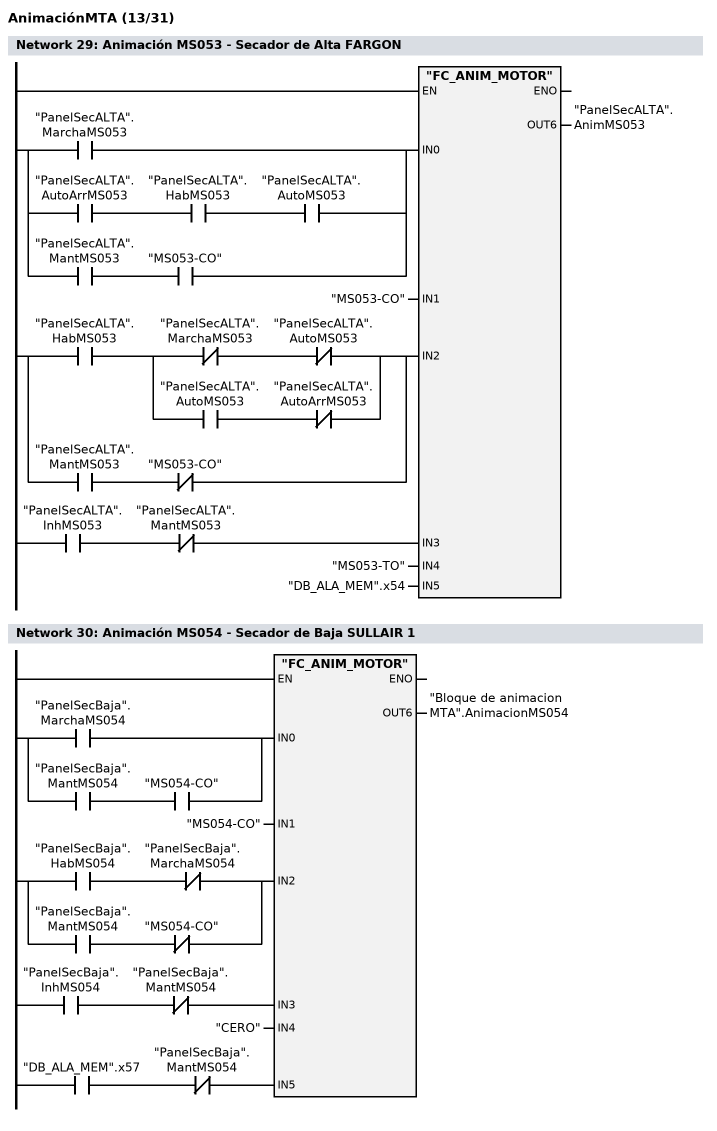
   RUNG wire#powerrail
      "FC_ANIM_MOTOR"(IN0 := wire#w1, IN2 := wire#w3, IN3 := wire#w4, IN1 := "MS053-CO", IN4 := "MS053-TO", IN5 := "DB_ALA_MEM".x54, OUT6 => "PanelSecALTA".AnimMS053)
   END_RUNG
   RUNG wire#powerrail
      Contact( "PanelSecALTA".MarchaMS053 )
   END_RUNG wire#w1
   RUNG wire#powerrail
      Contact( "PanelSecALTA".AutoArrMS053 )
      Contact( "PanelSecALTA".HabMS053 )
      Contact( "PanelSecALTA".AutoMS053 )
   END_RUNG wire#w1
   RUNG wire#powerrail
      Contact( "PanelSecALTA".MantMS053 )
      Contact( "MS053-CO" )
   END_RUNG wire#w1
   RUNG wire#powerrail
      Contact( "PanelSecALTA".HabMS053 )
      wire#w2
      I_Contact( "PanelSecALTA".MarchaMS053 )
      I_Contact( "PanelSecALTA".AutoMS053 )
   END_RUNG wire#w3
   RUNG wire#w2
      Contact( "PanelSecALTA".AutoMS053 )
      I_Contact( "PanelSecALTA".AutoArrMS053 )
   END_RUNG wire#w3
   RUNG wire#powerrail
      Contact( "PanelSecALTA".MantMS053 )
      I_Contact( "MS053-CO" )
   END_RUNG wire#w3
   RUNG wire#powerrail
      Contact( "PanelSecALTA".InhMS053 )
      I_Contact( "PanelSecALTA".MantMS053 )
   END_RUNG wire#w4
   // the same network as SCL:
   "FC_ANIM_MOTOR"(IN0 := "PanelSecALTA".MarchaMS053 OR ("PanelSecALTA".AutoArrMS053 AND "PanelSecALTA".HabMS053 AND "PanelSecALTA".AutoMS053) OR ("PanelSecALTA".MantMS053 AND "MS053-CO"),
                   IN1 := "MS053-CO",
                   IN2 := ("PanelSecALTA".HabMS053 AND ((NOT "PanelSecALTA".MarchaMS053 AND NOT "PanelSecALTA".AutoMS053) OR ("PanelSecALTA".AutoMS053 AND NOT "PanelSecALTA".AutoArrMS053))) OR ("PanelSecALTA".MantMS053 AND NOT "MS053-CO"),
                   IN3 := "PanelSecALTA".InhMS053 AND NOT "PanelSecALTA".MantMS053,
                   IN4 := "MS053-TO",
                   IN5 := "DB_ALA_MEM".x54,
                   OUT6 => "PanelSecALTA".AnimMS053);
END_REGION

REGION Network 30: Animación MS054 - Secador de Baja SULLAIR 1
   RUNG wire#powerrail
      "FC_ANIM_MOTOR"(IN0 := wire#w1, IN2 := wire#w2, IN3 := wire#w3, IN5 := wire#w4, IN1 := "MS054-CO", IN4 := "CERO", OUT6 => "Bloque de animacion MTA".AnimacionMS054)
   END_RUNG
   RUNG wire#powerrail
      Contact( "PanelSecBaja".MarchaMS054 )
   END_RUNG wire#w1
   RUNG wire#powerrail
      Contact( "PanelSecBaja".MantMS054 )
      Contact( "MS054-CO" )
   END_RUNG wire#w1
   RUNG wire#powerrail
      Contact( "PanelSecBaja".HabMS054 )
      I_Contact( "PanelSecBaja".MarchaMS054 )
   END_RUNG wire#w2
   RUNG wire#powerrail
      Contact( "PanelSecBaja".MantMS054 )
      I_Contact( "MS054-CO" )
   END_RUNG wire#w2
   RUNG wire#powerrail
      Contact( "PanelSecBaja".InhMS054 )
      I_Contact( "PanelSecBaja".MantMS054 )
   END_RUNG wire#w3
   RUNG wire#powerrail
      Contact( "DB_ALA_MEM".x57 )
      I_Contact( "PanelSecBaja".MantMS054 )
   END_RUNG wire#w4
   // the same network as SCL:
   "FC_ANIM_MOTOR"(IN0 := "PanelSecBaja".MarchaMS054 OR ("PanelSecBaja".MantMS054 AND "MS054-CO"),
                   IN1 := "MS054-CO",
                   IN2 := ("PanelSecBaja".HabMS054 AND NOT "PanelSecBaja".MarchaMS054) OR ("PanelSecBaja".MantMS054 AND NOT "MS054-CO"),
                   IN3 := "PanelSecBaja".InhMS054 AND NOT "PanelSecBaja".MantMS054,
                   IN4 := "CERO",
                   IN5 := "DB_ALA_MEM".x57 AND NOT "PanelSecBaja".MantMS054,
                   OUT6 => "Bloque de animacion MTA".AnimacionMS054);
END_REGION

REGION Network 31: Animación MS055 - Secador de Baja SULLAIR 2
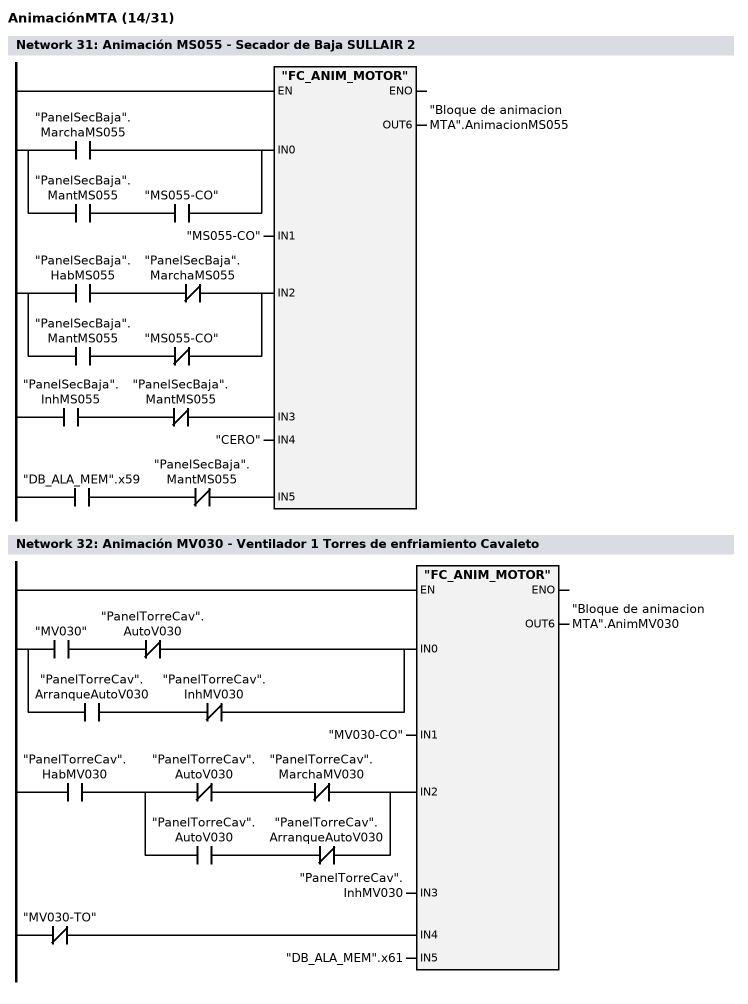
   RUNG wire#powerrail
      "FC_ANIM_MOTOR"(IN0 := wire#w1, IN2 := wire#w2, IN3 := wire#w3, IN5 := wire#w4, IN1 := "MS055-CO", IN4 := "CERO", OUT6 => "Bloque de animacion MTA".AnimacionMS055)
   END_RUNG
   RUNG wire#powerrail
      Contact( "PanelSecBaja".MarchaMS055 )
   END_RUNG wire#w1
   RUNG wire#powerrail
      Contact( "PanelSecBaja".MantMS055 )
      Contact( "MS055-CO" )
   END_RUNG wire#w1
   RUNG wire#powerrail
      Contact( "PanelSecBaja".HabMS055 )
      I_Contact( "PanelSecBaja".MarchaMS055 )
   END_RUNG wire#w2
   RUNG wire#powerrail
      Contact( "PanelSecBaja".MantMS055 )
      I_Contact( "MS055-CO" )
   END_RUNG wire#w2
   RUNG wire#powerrail
      Contact( "PanelSecBaja".InhMS055 )
      I_Contact( "PanelSecBaja".MantMS055 )
   END_RUNG wire#w3
   RUNG wire#powerrail
      Contact( "DB_ALA_MEM".x59 )
      I_Contact( "PanelSecBaja".MantMS055 )
   END_RUNG wire#w4
   // the same network as SCL:
   "FC_ANIM_MOTOR"(IN0 := "PanelSecBaja".MarchaMS055 OR ("PanelSecBaja".MantMS055 AND "MS055-CO"),
                   IN1 := "MS055-CO",
                   IN2 := ("PanelSecBaja".HabMS055 AND NOT "PanelSecBaja".MarchaMS055) OR ("PanelSecBaja".MantMS055 AND NOT "MS055-CO"),
                   IN3 := "PanelSecBaja".InhMS055 AND NOT "PanelSecBaja".MantMS055,
                   IN4 := "CERO",
                   IN5 := "DB_ALA_MEM".x59 AND NOT "PanelSecBaja".MantMS055,
                   OUT6 => "Bloque de animacion MTA".AnimacionMS055);
END_REGION

REGION Network 32: Animación MV030 - Ventilador 1 Torres de enfriamiento Cavaleto
   RUNG wire#powerrail
      "FC_ANIM_MOTOR"(IN0 := wire#w1, IN2 := wire#w3, IN4 := wire#w4, IN1 := "MV030-CO", IN3 := "PanelTorreCav".InhMV030, IN5 := "DB_ALA_MEM".x61, OUT6 => "Bloque de animacion MTA".AnimMV030)
   END_RUNG
   RUNG wire#powerrail
      Contact( "MV030" )
      I_Contact( "PanelTorreCav".AutoV030 )
   END_RUNG wire#w1
   RUNG wire#powerrail
      Contact( "PanelTorreCav".ArranqueAutoV030 )
      I_Contact( "PanelTorreCav".InhMV030 )
   END_RUNG wire#w1
   RUNG wire#powerrail
      Contact( "PanelTorreCav".HabMV030 )
      wire#w2
      I_Contact( "PanelTorreCav".AutoV030 )
      I_Contact( "PanelTorreCav".MarchaMV030 )
   END_RUNG wire#w3
   RUNG wire#w2
      Contact( "PanelTorreCav".AutoV030 )
      I_Contact( "PanelTorreCav".ArranqueAutoV030 )
   END_RUNG wire#w3
   RUNG wire#powerrail
      I_Contact( "MV030-TO" )
   END_RUNG wire#w4
   // the same network as SCL:
   "FC_ANIM_MOTOR"(IN0 := ("MV030" AND NOT "PanelTorreCav".AutoV030) OR ("PanelTorreCav".ArranqueAutoV030 AND NOT "PanelTorreCav".InhMV030),
                   IN1 := "MV030-CO",
                   IN2 := "PanelTorreCav".HabMV030 AND ((NOT "PanelTorreCav".AutoV030 AND NOT "PanelTorreCav".MarchaMV030) OR ("PanelTorreCav".AutoV030 AND NOT "PanelTorreCav".ArranqueAutoV030)),
                   IN3 := "PanelTorreCav".InhMV030,
                   IN4 := NOT "MV030-TO",
                   IN5 := "DB_ALA_MEM".x61,
                   OUT6 => "Bloque de animacion MTA".AnimMV030);
END_REGION

REGION Network 33: Animación MV031 - Ventilador 2 Torres de enfriamiento Cavaleto
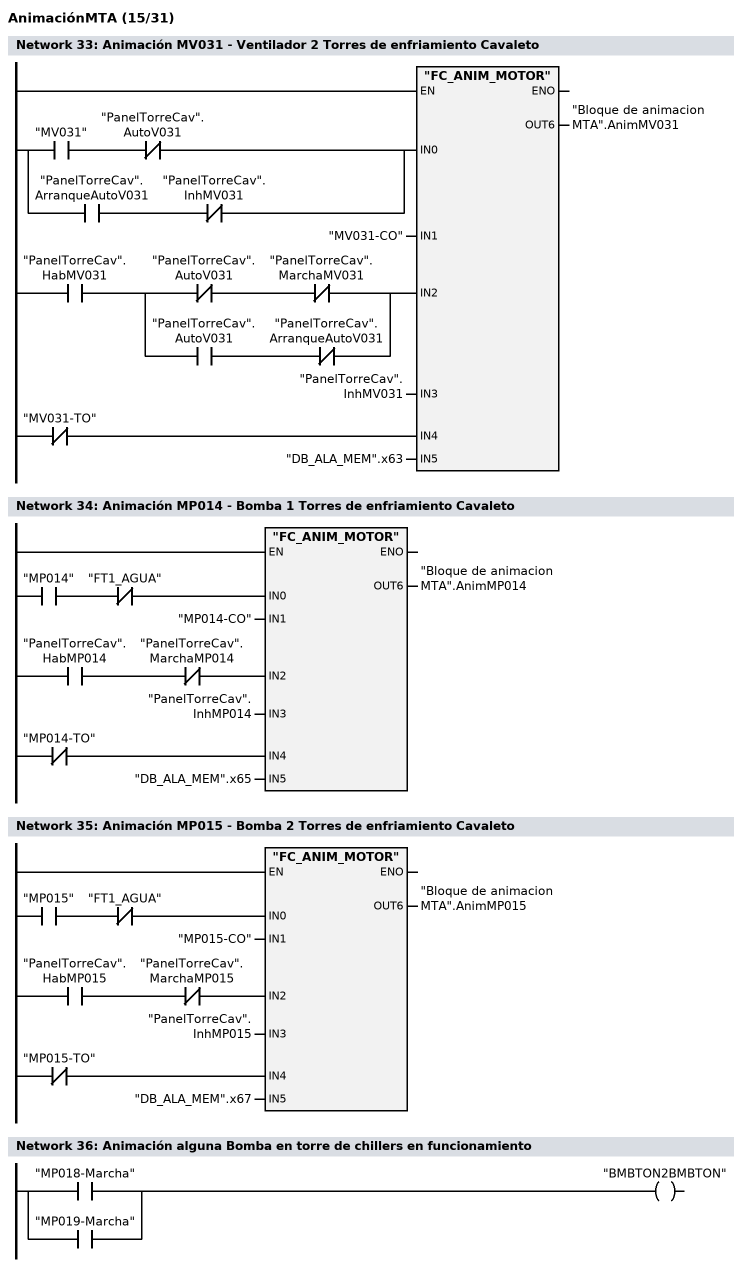
   RUNG wire#powerrail
      "FC_ANIM_MOTOR"(IN0 := wire#w1, IN2 := wire#w3, IN4 := wire#w4, IN1 := "MV031-CO", IN3 := "PanelTorreCav".InhMV031, IN5 := "DB_ALA_MEM".x63, OUT6 => "Bloque de animacion MTA".AnimMV031)
   END_RUNG
   RUNG wire#powerrail
      Contact( "MV031" )
      I_Contact( "PanelTorreCav".AutoV031 )
   END_RUNG wire#w1
   RUNG wire#powerrail
      Contact( "PanelTorreCav".ArranqueAutoV031 )
      I_Contact( "PanelTorreCav".InhMV031 )
   END_RUNG wire#w1
   RUNG wire#powerrail
      Contact( "PanelTorreCav".HabMV031 )
      wire#w2
      I_Contact( "PanelTorreCav".AutoV031 )
      I_Contact( "PanelTorreCav".MarchaMV031 )
   END_RUNG wire#w3
   RUNG wire#w2
      Contact( "PanelTorreCav".AutoV031 )
      I_Contact( "PanelTorreCav".ArranqueAutoV031 )
   END_RUNG wire#w3
   RUNG wire#powerrail
      I_Contact( "MV031-TO" )
   END_RUNG wire#w4
   // the same network as SCL:
   "FC_ANIM_MOTOR"(IN0 := ("MV031" AND NOT "PanelTorreCav".AutoV031) OR ("PanelTorreCav".ArranqueAutoV031 AND NOT "PanelTorreCav".InhMV031),
                   IN1 := "MV031-CO",
                   IN2 := "PanelTorreCav".HabMV031 AND ((NOT "PanelTorreCav".AutoV031 AND NOT "PanelTorreCav".MarchaMV031) OR ("PanelTorreCav".AutoV031 AND NOT "PanelTorreCav".ArranqueAutoV031)),
                   IN3 := "PanelTorreCav".InhMV031,
                   IN4 := NOT "MV031-TO",
                   IN5 := "DB_ALA_MEM".x63,
                   OUT6 => "Bloque de animacion MTA".AnimMV031);
END_REGION

REGION Network 34: Animación MP014 - Bomba 1 Torres de enfriamiento Cavaleto
   RUNG wire#powerrail
      "FC_ANIM_MOTOR"(IN0 := wire#w1, IN2 := wire#w2, IN4 := wire#w3, IN1 := "MP014-CO", IN3 := "PanelTorreCav".InhMP014, IN5 := "DB_ALA_MEM".x65, OUT6 => "Bloque de animacion MTA".AnimMP014)
   END_RUNG
   RUNG wire#powerrail
      Contact( "MP014" )
      I_Contact( "FT1_AGUA" )
   END_RUNG wire#w1
   RUNG wire#powerrail
      Contact( "PanelTorreCav".HabMP014 )
      I_Contact( "PanelTorreCav".MarchaMP014 )
   END_RUNG wire#w2
   RUNG wire#powerrail
      I_Contact( "MP014-TO" )
   END_RUNG wire#w3
   // the same network as SCL:
   "FC_ANIM_MOTOR"(IN0 := "MP014" AND NOT "FT1_AGUA",
                   IN1 := "MP014-CO",
                   IN2 := "PanelTorreCav".HabMP014 AND NOT "PanelTorreCav".MarchaMP014,
                   IN3 := "PanelTorreCav".InhMP014,
                   IN4 := NOT "MP014-TO",
                   IN5 := "DB_ALA_MEM".x65,
                   OUT6 => "Bloque de animacion MTA".AnimMP014);
END_REGION

REGION Network 35: Animación MP015 - Bomba 2 Torres de enfriamiento Cavaleto
   RUNG wire#powerrail
      "FC_ANIM_MOTOR"(IN0 := wire#w1, IN2 := wire#w2, IN4 := wire#w3, IN1 := "MP015-CO", IN3 := "PanelTorreCav".InhMP015, IN5 := "DB_ALA_MEM".x67, OUT6 => "Bloque de animacion MTA".AnimMP015)
   END_RUNG
   RUNG wire#powerrail
      Contact( "MP015" )
      I_Contact( "FT1_AGUA" )
   END_RUNG wire#w1
   RUNG wire#powerrail
      Contact( "PanelTorreCav".HabMP015 )
      I_Contact( "PanelTorreCav".MarchaMP015 )
   END_RUNG wire#w2
   RUNG wire#powerrail
      I_Contact( "MP015-TO" )
   END_RUNG wire#w3
   // the same network as SCL:
   "FC_ANIM_MOTOR"(IN0 := "MP015" AND NOT "FT1_AGUA",
                   IN1 := "MP015-CO",
                   IN2 := "PanelTorreCav".HabMP015 AND NOT "PanelTorreCav".MarchaMP015,
                   IN3 := "PanelTorreCav".InhMP015,
                   IN4 := NOT "MP015-TO",
                   IN5 := "DB_ALA_MEM".x67,
                   OUT6 => "Bloque de animacion MTA".AnimMP015);
END_REGION

REGION Network 36: Animación alguna Bomba en torre de chillers en funcionamiento
   RUNG wire#powerrail
      Contact( "MP018-Marcha" )
      wire#w1
      Coil( "BMBTON2BMBTON" )
   END_RUNG
   RUNG wire#powerrail
      Contact( "MP019-Marcha" )
   END_RUNG wire#w1
   // the same network as SCL:
   "BMBTON2BMBTON" := "MP018-Marcha" OR "MP019-Marcha";
END_REGION

REGION Network 37: Animación alguna Bomba en torre de cavaleto en funcionamiento
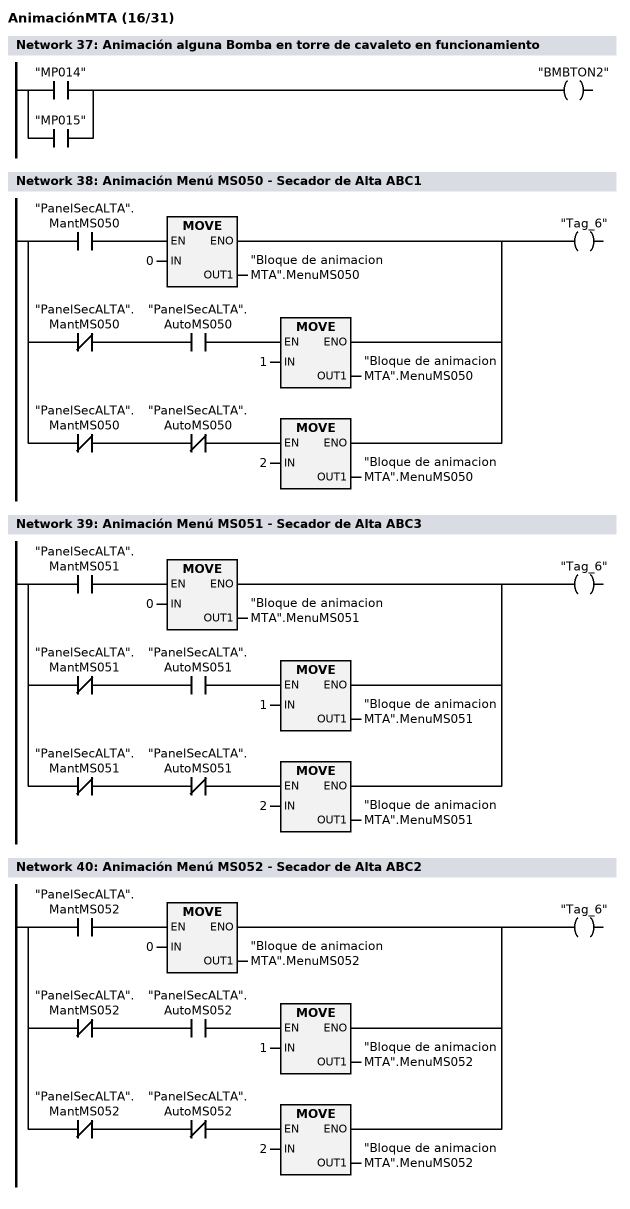
   RUNG wire#powerrail
      Contact( "MP014" )
      wire#w1
      Coil( "BMBTON2" )
   END_RUNG
   RUNG wire#powerrail
      Contact( "MP015" )
   END_RUNG wire#w1
   // the same network as SCL:
   "BMBTON2" := "MP014" OR "MP015";
END_REGION

REGION Network 38: Animación Menú MS050 - Secador de Alta ABC1
   RUNG wire#powerrail
      Contact( "PanelSecALTA".MantMS050 )
      { S7_GenerateENO := "TRUE" } Move(in := 0, out1 => "Bloque de animacion MTA".MenuMS050)
      wire#w1
      Coil( "Tag_6" )
   END_RUNG
   RUNG wire#powerrail
      I_Contact( "PanelSecALTA".MantMS050 )
      Contact( "PanelSecALTA".AutoMS050 )
      { S7_GenerateENO := "TRUE" } Move(in := 1, out1 => "Bloque de animacion MTA".MenuMS050)
   END_RUNG wire#w1
   RUNG wire#powerrail
      I_Contact( "PanelSecALTA".MantMS050 )
      I_Contact( "PanelSecALTA".AutoMS050 )
      { S7_GenerateENO := "TRUE" } Move(in := 2, out1 => "Bloque de animacion MTA".MenuMS050)
   END_RUNG wire#w1
   // the same network as SCL:
   // ENO of a box is taken as its EN; it also drops when the box reports an error
   IF "PanelSecALTA".MantMS050 THEN "Bloque de animacion MTA".MenuMS050 := 0; END_IF;
   #_w1 := NOT "PanelSecALTA".MantMS050 AND "PanelSecALTA".AutoMS050;
   IF #_w1 THEN "Bloque de animacion MTA".MenuMS050 := 1; END_IF;
   #_w2 := NOT "PanelSecALTA".MantMS050 AND NOT "PanelSecALTA".AutoMS050;
   IF #_w2 THEN "Bloque de animacion MTA".MenuMS050 := 2; END_IF;
   "Tag_6" := "PanelSecALTA".MantMS050 OR #_w1 OR #_w2;
END_REGION

REGION Network 39: Animación Menú MS051 - Secador de Alta ABC3
   RUNG wire#powerrail
      Contact( "PanelSecALTA".MantMS051 )
      { S7_GenerateENO := "TRUE" } Move(in := 0, out1 => "Bloque de animacion MTA".MenuMS051)
      wire#w1
      Coil( "Tag_6" )
   END_RUNG
   RUNG wire#powerrail
      I_Contact( "PanelSecALTA".MantMS051 )
      Contact( "PanelSecALTA".AutoMS051 )
      { S7_GenerateENO := "TRUE" } Move(in := 1, out1 => "Bloque de animacion MTA".MenuMS051)
   END_RUNG wire#w1
   RUNG wire#powerrail
      I_Contact( "PanelSecALTA".MantMS051 )
      I_Contact( "PanelSecALTA".AutoMS051 )
      { S7_GenerateENO := "TRUE" } Move(in := 2, out1 => "Bloque de animacion MTA".MenuMS051)
   END_RUNG wire#w1
   // the same network as SCL:
   // ENO of a box is taken as its EN; it also drops when the box reports an error
   IF "PanelSecALTA".MantMS051 THEN "Bloque de animacion MTA".MenuMS051 := 0; END_IF;
   #_w1 := NOT "PanelSecALTA".MantMS051 AND "PanelSecALTA".AutoMS051;
   IF #_w1 THEN "Bloque de animacion MTA".MenuMS051 := 1; END_IF;
   #_w2 := NOT "PanelSecALTA".MantMS051 AND NOT "PanelSecALTA".AutoMS051;
   IF #_w2 THEN "Bloque de animacion MTA".MenuMS051 := 2; END_IF;
   "Tag_6" := "PanelSecALTA".MantMS051 OR #_w1 OR #_w2;
END_REGION

REGION Network 40: Animación Menú MS052 - Secador de Alta ABC2
   RUNG wire#powerrail
      Contact( "PanelSecALTA".MantMS052 )
      { S7_GenerateENO := "TRUE" } Move(in := 0, out1 => "Bloque de animacion MTA".MenuMS052)
      wire#w1
      Coil( "Tag_6" )
   END_RUNG
   RUNG wire#powerrail
      I_Contact( "PanelSecALTA".MantMS052 )
      Contact( "PanelSecALTA".AutoMS052 )
      { S7_GenerateENO := "TRUE" } Move(in := 1, out1 => "Bloque de animacion MTA".MenuMS052)
   END_RUNG wire#w1
   RUNG wire#powerrail
      I_Contact( "PanelSecALTA".MantMS052 )
      I_Contact( "PanelSecALTA".AutoMS052 )
      { S7_GenerateENO := "TRUE" } Move(in := 2, out1 => "Bloque de animacion MTA".MenuMS052)
   END_RUNG wire#w1
   // the same network as SCL:
   // ENO of a box is taken as its EN; it also drops when the box reports an error
   IF "PanelSecALTA".MantMS052 THEN "Bloque de animacion MTA".MenuMS052 := 0; END_IF;
   #_w1 := NOT "PanelSecALTA".MantMS052 AND "PanelSecALTA".AutoMS052;
   IF #_w1 THEN "Bloque de animacion MTA".MenuMS052 := 1; END_IF;
   #_w2 := NOT "PanelSecALTA".MantMS052 AND NOT "PanelSecALTA".AutoMS052;
   IF #_w2 THEN "Bloque de animacion MTA".MenuMS052 := 2; END_IF;
   "Tag_6" := "PanelSecALTA".MantMS052 OR #_w1 OR #_w2;
END_REGION

REGION Network 41: Animación Menú MS053 - Secador de Alta FARGON
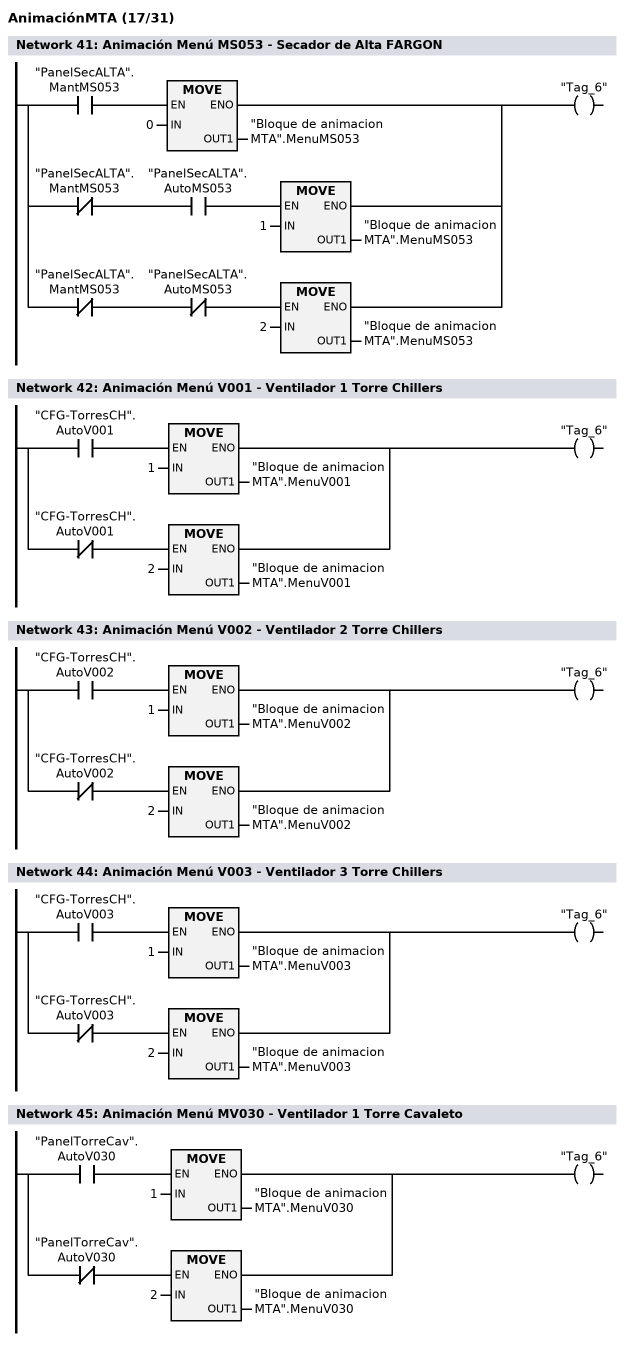
   RUNG wire#powerrail
      Contact( "PanelSecALTA".MantMS053 )
      { S7_GenerateENO := "TRUE" } Move(in := 0, out1 => "Bloque de animacion MTA".MenuMS053)
      wire#w1
      Coil( "Tag_6" )
   END_RUNG
   RUNG wire#powerrail
      I_Contact( "PanelSecALTA".MantMS053 )
      Contact( "PanelSecALTA".AutoMS053 )
      { S7_GenerateENO := "TRUE" } Move(in := 1, out1 => "Bloque de animacion MTA".MenuMS053)
   END_RUNG wire#w1
   RUNG wire#powerrail
      I_Contact( "PanelSecALTA".MantMS053 )
      I_Contact( "PanelSecALTA".AutoMS053 )
      { S7_GenerateENO := "TRUE" } Move(in := 2, out1 => "Bloque de animacion MTA".MenuMS053)
   END_RUNG wire#w1
   // the same network as SCL:
   // ENO of a box is taken as its EN; it also drops when the box reports an error
   IF "PanelSecALTA".MantMS053 THEN "Bloque de animacion MTA".MenuMS053 := 0; END_IF;
   #_w1 := NOT "PanelSecALTA".MantMS053 AND "PanelSecALTA".AutoMS053;
   IF #_w1 THEN "Bloque de animacion MTA".MenuMS053 := 1; END_IF;
   #_w2 := NOT "PanelSecALTA".MantMS053 AND NOT "PanelSecALTA".AutoMS053;
   IF #_w2 THEN "Bloque de animacion MTA".MenuMS053 := 2; END_IF;
   "Tag_6" := "PanelSecALTA".MantMS053 OR #_w1 OR #_w2;
END_REGION

REGION Network 42: Animación Menú V001 - Ventilador 1 Torre Chillers
   RUNG wire#powerrail
      Contact( "CFG-TorresCH".AutoV001 )
      { S7_GenerateENO := "TRUE" } Move(in := 1, out1 => "Bloque de animacion MTA".MenuV001)
      wire#w1
      Coil( "Tag_6" )
   END_RUNG
   RUNG wire#powerrail
      I_Contact( "CFG-TorresCH".AutoV001 )
      { S7_GenerateENO := "TRUE" } Move(in := 2, out1 => "Bloque de animacion MTA".MenuV001)
   END_RUNG wire#w1
   // the same network as SCL:
   // ENO of a box is taken as its EN; it also drops when the box reports an error
   IF "CFG-TorresCH".AutoV001 THEN "Bloque de animacion MTA".MenuV001 := 1; END_IF;
   #_w1 := NOT "CFG-TorresCH".AutoV001;
   IF #_w1 THEN "Bloque de animacion MTA".MenuV001 := 2; END_IF;
   "Tag_6" := "CFG-TorresCH".AutoV001 OR #_w1;
END_REGION

REGION Network 43: Animación Menú V002 - Ventilador 2 Torre Chillers
   RUNG wire#powerrail
      Contact( "CFG-TorresCH".AutoV002 )
      { S7_GenerateENO := "TRUE" } Move(in := 1, out1 => "Bloque de animacion MTA".MenuV002)
      wire#w1
      Coil( "Tag_6" )
   END_RUNG
   RUNG wire#powerrail
      I_Contact( "CFG-TorresCH".AutoV002 )
      { S7_GenerateENO := "TRUE" } Move(in := 2, out1 => "Bloque de animacion MTA".MenuV002)
   END_RUNG wire#w1
   // the same network as SCL:
   // ENO of a box is taken as its EN; it also drops when the box reports an error
   IF "CFG-TorresCH".AutoV002 THEN "Bloque de animacion MTA".MenuV002 := 1; END_IF;
   #_w1 := NOT "CFG-TorresCH".AutoV002;
   IF #_w1 THEN "Bloque de animacion MTA".MenuV002 := 2; END_IF;
   "Tag_6" := "CFG-TorresCH".AutoV002 OR #_w1;
END_REGION

REGION Network 44: Animación Menú V003 - Ventilador 3 Torre Chillers
   RUNG wire#powerrail
      Contact( "CFG-TorresCH".AutoV003 )
      { S7_GenerateENO := "TRUE" } Move(in := 1, out1 => "Bloque de animacion MTA".MenuV003)
      wire#w1
      Coil( "Tag_6" )
   END_RUNG
   RUNG wire#powerrail
      I_Contact( "CFG-TorresCH".AutoV003 )
      { S7_GenerateENO := "TRUE" } Move(in := 2, out1 => "Bloque de animacion MTA".MenuV003)
   END_RUNG wire#w1
   // the same network as SCL:
   // ENO of a box is taken as its EN; it also drops when the box reports an error
   IF "CFG-TorresCH".AutoV003 THEN "Bloque de animacion MTA".MenuV003 := 1; END_IF;
   #_w1 := NOT "CFG-TorresCH".AutoV003;
   IF #_w1 THEN "Bloque de animacion MTA".MenuV003 := 2; END_IF;
   "Tag_6" := "CFG-TorresCH".AutoV003 OR #_w1;
END_REGION

REGION Network 45: Animación Menú MV030 - Ventilador 1 Torre Cavaleto
   RUNG wire#powerrail
      Contact( "PanelTorreCav".AutoV030 )
      { S7_GenerateENO := "TRUE" } Move(in := 1, out1 => "Bloque de animacion MTA".MenuV030)
      wire#w1
      Coil( "Tag_6" )
   END_RUNG
   RUNG wire#powerrail
      I_Contact( "PanelTorreCav".AutoV030 )
      { S7_GenerateENO := "TRUE" } Move(in := 2, out1 => "Bloque de animacion MTA".MenuV030)
   END_RUNG wire#w1
   // the same network as SCL:
   // ENO of a box is taken as its EN; it also drops when the box reports an error
   IF "PanelTorreCav".AutoV030 THEN "Bloque de animacion MTA".MenuV030 := 1; END_IF;
   #_w1 := NOT "PanelTorreCav".AutoV030;
   IF #_w1 THEN "Bloque de animacion MTA".MenuV030 := 2; END_IF;
   "Tag_6" := "PanelTorreCav".AutoV030 OR #_w1;
END_REGION

REGION Network 46: Animación Menú MV031 - Ventilador 2 Torre Cavaleto
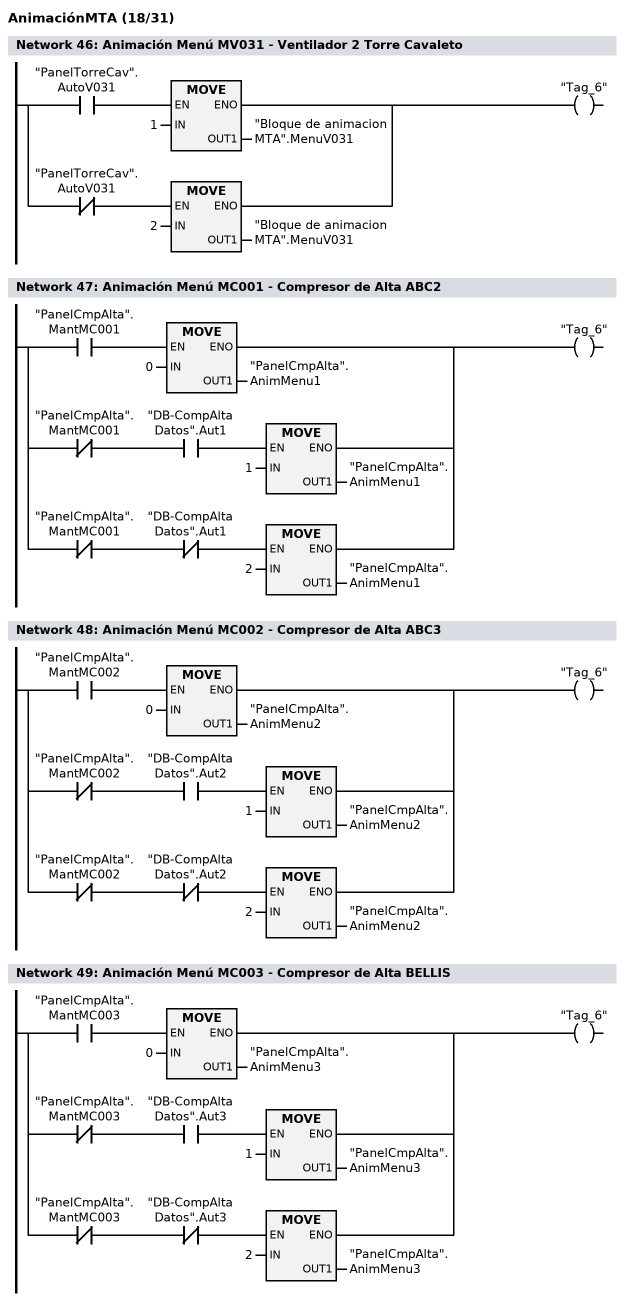
   RUNG wire#powerrail
      Contact( "PanelTorreCav".AutoV031 )
      { S7_GenerateENO := "TRUE" } Move(in := 1, out1 => "Bloque de animacion MTA".MenuV031)
      wire#w1
      Coil( "Tag_6" )
   END_RUNG
   RUNG wire#powerrail
      I_Contact( "PanelTorreCav".AutoV031 )
      { S7_GenerateENO := "TRUE" } Move(in := 2, out1 => "Bloque de animacion MTA".MenuV031)
   END_RUNG wire#w1
   // the same network as SCL:
   // ENO of a box is taken as its EN; it also drops when the box reports an error
   IF "PanelTorreCav".AutoV031 THEN "Bloque de animacion MTA".MenuV031 := 1; END_IF;
   #_w1 := NOT "PanelTorreCav".AutoV031;
   IF #_w1 THEN "Bloque de animacion MTA".MenuV031 := 2; END_IF;
   "Tag_6" := "PanelTorreCav".AutoV031 OR #_w1;
END_REGION

REGION Network 47: Animación Menú MC001 - Compresor de Alta ABC2
   RUNG wire#powerrail
      Contact( "PanelCmpAlta".MantMC001 )
      { S7_GenerateENO := "TRUE" } Move(in := 0, out1 => "PanelCmpAlta".AnimMenu1)
      wire#w1
      Coil( "Tag_6" )
   END_RUNG
   RUNG wire#powerrail
      I_Contact( "PanelCmpAlta".MantMC001 )
      Contact( "DB-CompAltaDatos".Aut1 )
      { S7_GenerateENO := "TRUE" } Move(in := 1, out1 => "PanelCmpAlta".AnimMenu1)
   END_RUNG wire#w1
   RUNG wire#powerrail
      I_Contact( "PanelCmpAlta".MantMC001 )
      I_Contact( "DB-CompAltaDatos".Aut1 )
      { S7_GenerateENO := "TRUE" } Move(in := 2, out1 => "PanelCmpAlta".AnimMenu1)
   END_RUNG wire#w1
   // the same network as SCL:
   // ENO of a box is taken as its EN; it also drops when the box reports an error
   IF "PanelCmpAlta".MantMC001 THEN "PanelCmpAlta".AnimMenu1 := 0; END_IF;
   #_w1 := NOT "PanelCmpAlta".MantMC001 AND "DB-CompAltaDatos".Aut1;
   IF #_w1 THEN "PanelCmpAlta".AnimMenu1 := 1; END_IF;
   #_w2 := NOT "PanelCmpAlta".MantMC001 AND NOT "DB-CompAltaDatos".Aut1;
   IF #_w2 THEN "PanelCmpAlta".AnimMenu1 := 2; END_IF;
   "Tag_6" := "PanelCmpAlta".MantMC001 OR #_w1 OR #_w2;
END_REGION

REGION Network 48: Animación Menú MC002 - Compresor de Alta ABC3
   RUNG wire#powerrail
      Contact( "PanelCmpAlta".MantMC002 )
      { S7_GenerateENO := "TRUE" } Move(in := 0, out1 => "PanelCmpAlta".AnimMenu2)
      wire#w1
      Coil( "Tag_6" )
   END_RUNG
   RUNG wire#powerrail
      I_Contact( "PanelCmpAlta".MantMC002 )
      Contact( "DB-CompAltaDatos".Aut2 )
      { S7_GenerateENO := "TRUE" } Move(in := 1, out1 => "PanelCmpAlta".AnimMenu2)
   END_RUNG wire#w1
   RUNG wire#powerrail
      I_Contact( "PanelCmpAlta".MantMC002 )
      I_Contact( "DB-CompAltaDatos".Aut2 )
      { S7_GenerateENO := "TRUE" } Move(in := 2, out1 => "PanelCmpAlta".AnimMenu2)
   END_RUNG wire#w1
   // the same network as SCL:
   // ENO of a box is taken as its EN; it also drops when the box reports an error
   IF "PanelCmpAlta".MantMC002 THEN "PanelCmpAlta".AnimMenu2 := 0; END_IF;
   #_w1 := NOT "PanelCmpAlta".MantMC002 AND "DB-CompAltaDatos".Aut2;
   IF #_w1 THEN "PanelCmpAlta".AnimMenu2 := 1; END_IF;
   #_w2 := NOT "PanelCmpAlta".MantMC002 AND NOT "DB-CompAltaDatos".Aut2;
   IF #_w2 THEN "PanelCmpAlta".AnimMenu2 := 2; END_IF;
   "Tag_6" := "PanelCmpAlta".MantMC002 OR #_w1 OR #_w2;
END_REGION

REGION Network 49: Animación Menú MC003 - Compresor de Alta BELLIS
   RUNG wire#powerrail
      Contact( "PanelCmpAlta".MantMC003 )
      { S7_GenerateENO := "TRUE" } Move(in := 0, out1 => "PanelCmpAlta".AnimMenu3)
      wire#w1
      Coil( "Tag_6" )
   END_RUNG
   RUNG wire#powerrail
      I_Contact( "PanelCmpAlta".MantMC003 )
      Contact( "DB-CompAltaDatos".Aut3 )
      { S7_GenerateENO := "TRUE" } Move(in := 1, out1 => "PanelCmpAlta".AnimMenu3)
   END_RUNG wire#w1
   RUNG wire#powerrail
      I_Contact( "PanelCmpAlta".MantMC003 )
      I_Contact( "DB-CompAltaDatos".Aut3 )
      { S7_GenerateENO := "TRUE" } Move(in := 2, out1 => "PanelCmpAlta".AnimMenu3)
   END_RUNG wire#w1
   // the same network as SCL:
   // ENO of a box is taken as its EN; it also drops when the box reports an error
   IF "PanelCmpAlta".MantMC003 THEN "PanelCmpAlta".AnimMenu3 := 0; END_IF;
   #_w1 := NOT "PanelCmpAlta".MantMC003 AND "DB-CompAltaDatos".Aut3;
   IF #_w1 THEN "PanelCmpAlta".AnimMenu3 := 1; END_IF;
   #_w2 := NOT "PanelCmpAlta".MantMC003 AND NOT "DB-CompAltaDatos".Aut3;
   IF #_w2 THEN "PanelCmpAlta".AnimMenu3 := 2; END_IF;
   "Tag_6" := "PanelCmpAlta".MantMC003 OR #_w1 OR #_w2;
END_REGION

REGION Network 50: Animación Menú MC004 - Compresor de Alta ABC4
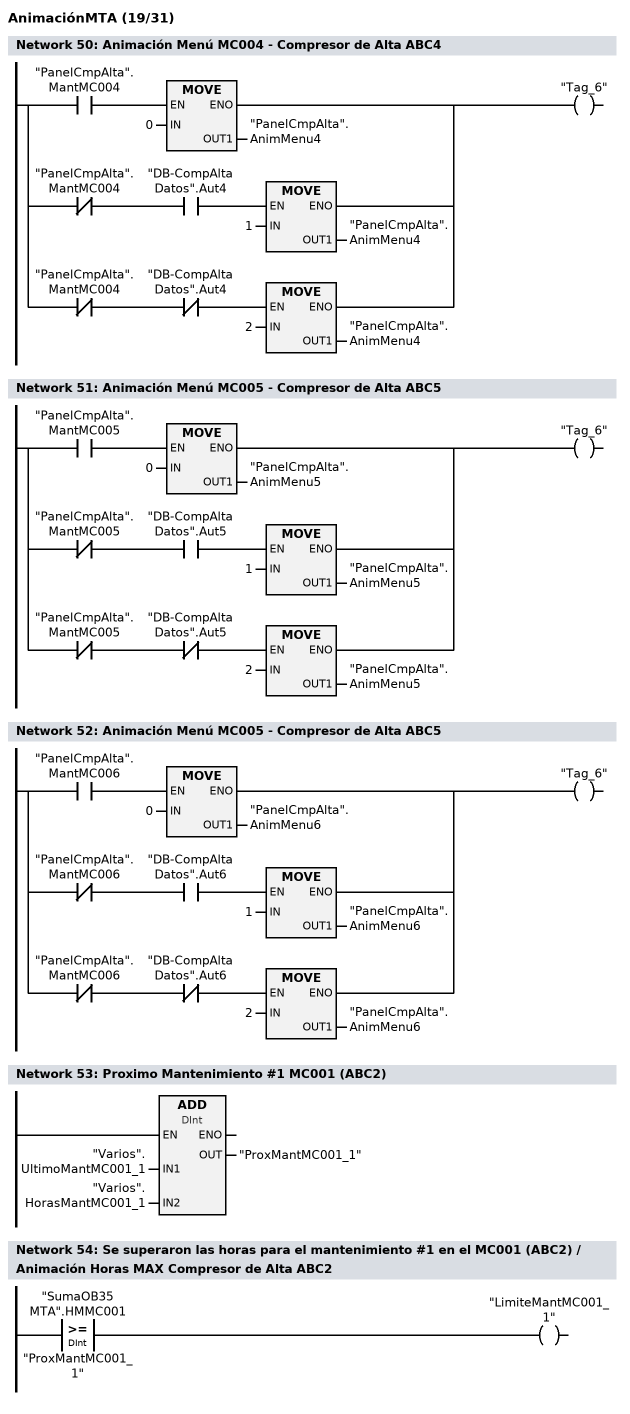
   RUNG wire#powerrail
      Contact( "PanelCmpAlta".MantMC004 )
      { S7_GenerateENO := "TRUE" } Move(in := 0, out1 => "PanelCmpAlta".AnimMenu4)
      wire#w1
      Coil( "Tag_6" )
   END_RUNG
   RUNG wire#powerrail
      I_Contact( "PanelCmpAlta".MantMC004 )
      Contact( "DB-CompAltaDatos".Aut4 )
      { S7_GenerateENO := "TRUE" } Move(in := 1, out1 => "PanelCmpAlta".AnimMenu4)
   END_RUNG wire#w1
   RUNG wire#powerrail
      I_Contact( "PanelCmpAlta".MantMC004 )
      I_Contact( "DB-CompAltaDatos".Aut4 )
      { S7_GenerateENO := "TRUE" } Move(in := 2, out1 => "PanelCmpAlta".AnimMenu4)
   END_RUNG wire#w1
   // the same network as SCL:
   // ENO of a box is taken as its EN; it also drops when the box reports an error
   IF "PanelCmpAlta".MantMC004 THEN "PanelCmpAlta".AnimMenu4 := 0; END_IF;
   #_w1 := NOT "PanelCmpAlta".MantMC004 AND "DB-CompAltaDatos".Aut4;
   IF #_w1 THEN "PanelCmpAlta".AnimMenu4 := 1; END_IF;
   #_w2 := NOT "PanelCmpAlta".MantMC004 AND NOT "DB-CompAltaDatos".Aut4;
   IF #_w2 THEN "PanelCmpAlta".AnimMenu4 := 2; END_IF;
   "Tag_6" := "PanelCmpAlta".MantMC004 OR #_w1 OR #_w2;
END_REGION

REGION Network 51: Animación Menú MC005 - Compresor de Alta ABC5
   RUNG wire#powerrail
      Contact( "PanelCmpAlta".MantMC005 )
      { S7_GenerateENO := "TRUE" } Move(in := 0, out1 => "PanelCmpAlta".AnimMenu5)
      wire#w1
      Coil( "Tag_6" )
   END_RUNG
   RUNG wire#powerrail
      I_Contact( "PanelCmpAlta".MantMC005 )
      Contact( "DB-CompAltaDatos".Aut5 )
      { S7_GenerateENO := "TRUE" } Move(in := 1, out1 => "PanelCmpAlta".AnimMenu5)
   END_RUNG wire#w1
   RUNG wire#powerrail
      I_Contact( "PanelCmpAlta".MantMC005 )
      I_Contact( "DB-CompAltaDatos".Aut5 )
      { S7_GenerateENO := "TRUE" } Move(in := 2, out1 => "PanelCmpAlta".AnimMenu5)
   END_RUNG wire#w1
   // the same network as SCL:
   // ENO of a box is taken as its EN; it also drops when the box reports an error
   IF "PanelCmpAlta".MantMC005 THEN "PanelCmpAlta".AnimMenu5 := 0; END_IF;
   #_w1 := NOT "PanelCmpAlta".MantMC005 AND "DB-CompAltaDatos".Aut5;
   IF #_w1 THEN "PanelCmpAlta".AnimMenu5 := 1; END_IF;
   #_w2 := NOT "PanelCmpAlta".MantMC005 AND NOT "DB-CompAltaDatos".Aut5;
   IF #_w2 THEN "PanelCmpAlta".AnimMenu5 := 2; END_IF;
   "Tag_6" := "PanelCmpAlta".MantMC005 OR #_w1 OR #_w2;
END_REGION

REGION Network 52: Animación Menú MC005 - Compresor de Alta ABC5
   RUNG wire#powerrail
      Contact( "PanelCmpAlta".MantMC006 )
      { S7_GenerateENO := "TRUE" } Move(in := 0, out1 => "PanelCmpAlta".AnimMenu6)
      wire#w1
      Coil( "Tag_6" )
   END_RUNG
   RUNG wire#powerrail
      I_Contact( "PanelCmpAlta".MantMC006 )
      Contact( "DB-CompAltaDatos".Aut6 )
      { S7_GenerateENO := "TRUE" } Move(in := 1, out1 => "PanelCmpAlta".AnimMenu6)
   END_RUNG wire#w1
   RUNG wire#powerrail
      I_Contact( "PanelCmpAlta".MantMC006 )
      I_Contact( "DB-CompAltaDatos".Aut6 )
      { S7_GenerateENO := "TRUE" } Move(in := 2, out1 => "PanelCmpAlta".AnimMenu6)
   END_RUNG wire#w1
   // the same network as SCL:
   // ENO of a box is taken as its EN; it also drops when the box reports an error
   IF "PanelCmpAlta".MantMC006 THEN "PanelCmpAlta".AnimMenu6 := 0; END_IF;
   #_w1 := NOT "PanelCmpAlta".MantMC006 AND "DB-CompAltaDatos".Aut6;
   IF #_w1 THEN "PanelCmpAlta".AnimMenu6 := 1; END_IF;
   #_w2 := NOT "PanelCmpAlta".MantMC006 AND NOT "DB-CompAltaDatos".Aut6;
   IF #_w2 THEN "PanelCmpAlta".AnimMenu6 := 2; END_IF;
   "Tag_6" := "PanelCmpAlta".MantMC006 OR #_w1 OR #_w2;
END_REGION

REGION Network 53: Proximo Mantenimiento #1 MC001 (ABC2)
   RUNG wire#powerrail
      { S7_Templates := "SrcType := DInt"; S7_GenerateENO := "TRUE" } Add(in1 := "Varios".UltimoMantMC001_1, in2 := "Varios".HorasMantMC001_1, out => "ProxMantMC001_1")
   END_RUNG
   // the same network as SCL:
   "ProxMantMC001_1" := "Varios".UltimoMantMC001_1 + "Varios".HorasMantMC001_1;
END_REGION

REGION Network 54: Se superaron las horas para el mantenimiento #1 en el MC001 (ABC2) / Animación Horas MAX Compresor de Alta ABC2
   RUNG wire#powerrail
      { S7_Templates := "SrcType := DInt" } GE_Contact(in1 := "SumaOB35 MTA".HMMC001, in2 := "ProxMantMC001_1")
      Coil( "LimiteMantMC001_1" )
   END_RUNG
   // the same network as SCL:
   "LimiteMantMC001_1" := "SumaOB35 MTA".HMMC001 >= "ProxMantMC001_1";
END_REGION

REGION Network 55: Proximo Mantenimiento #1 MC002 (ABC3)